   END_REGION

   REGION "CHANGE DETECTION"
       #old.btnParam := #btnParams;
       #old.kp8DI := #kp8DI;
       #old.logical := #retLogical.acutal;
       #old.physical := #btnPress;
   END_REGION

   REGION "OUTPUT"
       #kp8DQ := #colorMask;
       #physical := #retPhysical;
       #logical := #retLogical;
   END_REGION
END_FUNCTION_BLOCK

FUNCTION "KP8 Driver: HMI Emulator: Animation" : USInt   // FC26, SCL
{ S7_Optimized_Access := 'TRUE' }
VERSION : 0.1
   VAR_INPUT
      kp8Color : DWord;
      btnNumber : Int;
   END_VAR
   VAR_TEMP
      animate : USInt;
      blue : USInt;
      colorDWord : DWord;
      colorInt : DInt;
      green : USInt;
      off : USInt;
      red : USInt;
      white : USInt;
      yellow : USInt;
   END_VAR
   VAR CONSTANT
      blueMask : DInt := 16#0000_0100;
      btnMask : DInt := 16#0101_0100;
      greenMask : DInt := 16#0001_0000;
      offMask : DInt := 16#0000_0000;
      redMask : DInt := 16#0100_0000;
      whiteMask : DInt := 16#0101_0100;
      yellowMask : DInt := 16#0101_0000;
   END_VAR
BEGIN
   REGION "COPY TO LOCAL"
       #blue := "BLUE_LIGHT_BACKGROUND";
       #green := "GREEN_LIGHT_BACKGROUND";
       #off := "INVISIBLE";
       #red := "RED_LIGHT_BACKGROUND";
       #white := "WHITE_BACKGROUND";
       #yellow := "YELLOW_LIGHT_BACKGROUND";
   END_REGION

   REGION "ISOLATE BUTTON COLOR"
       #colorDWord := SHR_DWORD(IN := #kp8Color,N := INT_TO_ULINT(#btnNumber));
       #colorDWord := #colorDWord AND #btnMask;
       #colorInt := DWORD_TO_DINT(#colorDWord);
   END_REGION

   REGION "DETERMINE ANIMATION"
       CASE #colorInt OF
           #blueMask:
               #animate := #blue;
           #greenMask:
               #animate := #green;
           #redMask:
               #animate := #red;
           #whiteMask:
               #animate := #white;
           #yellowMask:
               #animate := #yellow;
           ELSE
               #animate := #off;
       END_CASE;
   END_REGION

   REGION "RETURN VALUE"
       #"KP8 Driver: HMI Emulator: Animation" := #animate;
   END_REGION
END_FUNCTION

FUNCTION "KP8 Driver: Group" : Void   // FC50, SCL
{ S7_Optimized_Access := 'TRUE' }
VERSION : 0.1
   VAR_INPUT
      btnNumber : Int;
      btnsParams : "KP8 Driver: Parameters: 8 Buttons";
   END_VAR
   VAR_IN_OUT
      logical : "KP8 Driver: Feedback Data";
   END_VAR
   VAR_TEMP
      pBtn : Int;
      retLogical : "KP8 Driver: Feedback Data";
      testGroup : Int;
      thisGroup : Int;
   END_VAR
BEGIN
   REGION "EXIT IF GROUP EQUALS 0"
       #thisGroup := #btnsParams.btn[#btnNumber].group;
       IF #thisGroup = 0 THEN
           RETURN;
       END_IF;
   END_REGION

   REGION "COPY TO LOCAL"
       #retLogical := #logical;
   END_REGION

   REGION "FOR EACH BUTTONS' PARAMETERS"
       FOR #pBtn := 0 TO 7 DO

           REGION "SKIP THE CURRENT BUTTON"
               IF #pBtn = #btnNumber THEN
                   GOTO NEXT;
               END_IF;
           END_REGION

           REGION "GROUP EXCLUSION"
               #testGroup := #btnsParams.btn[#pBtn].group;
               IF #testGroup = #thisGroup THEN
                   #retLogical.acutal.btn[#pBtn] := FALSE;
               END_IF;
           END_REGION

       NEXT:
           ;

       END_FOR;
   END_REGION

   REGION "OUTPUT"
       #logical := #retLogical;
   END_REGION
END_FUNCTION

FUNCTION "KP8 Driver: Toggle" : Void   // FC51, SCL
{ S7_Optimized_Access := 'TRUE' }
VERSION : 0.1
   VAR_INPUT
      signal : Bool;   // edge signal
   END_VAR
   VAR_IN_OUT
      state : Bool;   // logical button state
   END_VAR
BEGIN
   IF #signal THEN
       #state := NOT #state;
   END_IF;
END_FUNCTION

FUNCTION "KP8 Driver: Feedback" : Void   // FC52, SCL
{ S7_Optimized_Access := 'TRUE' }
VERSION : 0.1
   VAR_INPUT
      signal : Bool;
      oldSignal : Bool;
      btnNumber : Int;
   END_VAR
   VAR_IN_OUT
      feedback : "KP8 Driver: Feedback Data";
   END_VAR
   VAR_TEMP
      ret : "KP8 Driver: Feedback Data";
   END_VAR
BEGIN
   REGION "COPY TO LOCAL"
       #ret := #feedback;
       #ret.acutal.btn[#btnNumber] := #signal;
   END_REGION

   REGION "DEFAULT"
       #ret.rising.btn[#btnNumber] := FALSE;
       #ret.falling.btn[#btnNumber] := FALSE;
   END_REGION

   REGION "ON NEW INPUT"
       IF #signal <> #oldSignal THEN

           REGION "RISING EDGE"
               IF #signal AND NOT #oldSignal THEN
                   #ret.rising.btn[#btnNumber] := TRUE;
               END_IF;
           END_REGION

           REGION "FALLING EDGE"
               IF NOT #signal AND #oldSignal THEN
                   #ret.falling.btn[#btnNumber] := TRUE;
               END_IF;
           END_REGION

       END_IF;
   END_REGION


   REGION "OUTPUT"
       #feedback := #ret;
   END_REGION
END_FUNCTION

FUNCTION "KP8 Driver: State" : Void   // FC53, SCL
{ S7_Optimized_Access := 'TRUE' }
VERSION : 0.1
   VAR_INPUT
      press : "KP8 Driver: Feedback Data";
      btnNumber : Int;
      btnParams : "KP8 Driver: Parameters: 8 Buttons";
   END_VAR
   VAR_IN_OUT
      state : "KP8 Driver: Feedback Data";
   END_VAR
   VAR_TEMP
      pBtn : Int;
      retState : "KP8 Driver: Feedback Data";
   END_VAR
BEGIN
   REGION "RETURN ON INACTIVE BUTTON"
       IF NOT #btnParams.btn[#btnNumber].activate THEN
           RETURN;
       END_IF;
   END_REGION

   REGION "COPY TO LOCAL"
       #retState := #state;
   END_REGION

   REGION "MODE IS MOMENTARY"
       IF NOT #btnParams.btn[#btnNumber].mode THEN
           #retState.acutal.btn[#btnNumber] := #press.acutal.btn[#btnNumber];
       END_IF;
   END_REGION

   REGION "MAINTINED"
       IF #btnParams.btn[#btnNumber].mode THEN
           "KP8 Driver: Toggle"(signal := #press.rising.btn[#btnNumber],
                                state := #retState.acutal.btn[#btnNumber]);
       END_IF;
   END_REGION

   REGION "GROUP EXCLUSIVITY"
       IF #press.rising.btn[#btnNumber] THEN
           "KP8 Driver: Group"(btnNumber := #btnNumber,
                               btnsParams := #btnParams,
                               logical := #retState);
       END_IF;
   END_REGION

   REGION "OUTPUT"
       #state := #retState;
   END_REGION
END_FUNCTION

FUNCTION "KP8 Driver: Color" : Void   // FC54, SCL
{ S7_Optimized_Access := 'TRUE' }
VERSION : 0.1
   VAR_INPUT
      btnNum : Int;
      lblColor : String;   // 'red', 'green', 'blue', 'yellow', 'white', 'off'
   END_VAR
   VAR_IN_OUT
      btnColor : DWord;
   END_VAR
   VAR_TEMP
      btnMask : DWord;
      uColor : String;
      ret : DWord;
   END_VAR
   VAR CONSTANT
      btnMskRed : DWord := DWORD#16#0100_0000;
      btnMskGreen : DWord := DWORD#16#0001_0000;
      btnMskBlue : DWord := DWORD#16#0000_0100;
      btnMskYellow : DWord := DWORD#16#0101_0000;
      btnMskWhite : DWord := DWORD#16#0101_0100;
      btnMskOff : DWord := DWORD#16#FEFE_FEFF;
   END_VAR
BEGIN
   #ret := #btnColor;

   #ret := #ret AND ROL(IN := #btnMskOff,
                        N := INT_TO_UDINT(#btnNum));

   #uColor := #lblColor;
   "Upper"(#uColor);

   IF (#uColor = 'RED') THEN
       #btnMask := #btnMskRed;
   ELSIF (#uColor = 'GREEN') THEN
       #btnMask := #btnMskGreen;
   ELSIF (#uColor = 'BLUE') THEN
       #btnMask := #btnMskBlue;
   ELSIF (#uColor = 'YELLOW') THEN
       #btnMask := #btnMskYellow;
   ELSIF (#uColor = 'WHITE') THEN
       #btnMask := #btnMskWhite;
   ELSIF (#uColor = 'OFF') THEN
       ;
   END_IF;

   #ret := #ret OR SHL(IN := #btnMask,
                       N := INT_TO_UDINT(#btnNum));

   #btnColor := #ret;
END_FUNCTION

FUNCTION "KP8 Driver: HMI Emulator: Button Presses" : Word   // FC82, SCL
{ S7_Optimized_Access := 'TRUE' }
VERSION : 0.1
   VAR_INPUT
      pbs : DWord;
   END_VAR
   VAR_TEMP
      ret : Word;
   END_VAR
BEGIN
   #"KP8 Driver: HMI Emulator: Button Presses".%B1 := #pbs.%B0;
   #"KP8 Driver: HMI Emulator: Button Presses".%B0 := #pbs.%B1;
END_FUNCTION

// folder: Utilities

FUNCTION_BLOCK "Pulses: Button Collection"   // FB22, SCL
{ S7_Optimized_Access := 'TRUE' }
VERSION : 0.1
   VAR_INPUT
      btns : Variant;
   END_VAR
   VAR_IN_OUT
      pulses : Variant;
   END_VAR
   VAR
      old : Array[0..#u_bound] of Int;
   END_VAR
   VAR_TEMP
      eval : Array[0..#u_bound] of Int;
      i : Int;
      len_btns : UDInt;
      ret : Array[0..#u_bound] of Int;
      RET_VAL : Int;
   END_VAR
   VAR CONSTANT
      u_bound : Int := 999;
   END_VAR
BEGIN
   REGION "GET ARRAY LENGTH"
       #len_btns := CountOfElements(#btns);
   END_REGION


   REGION "COPY TO LOCAL"
       #RET_VAL := MOVE_BLK_VARIANT(SRC := #btns,
                                    COUNT := #len_btns,
                                    SRC_INDEX := 0,
                                    DEST_INDEX := 0,
                                    DEST => #eval);
   END_REGION


   REGION "CHECK FOR FALLING EDGE"
       FOR #i := 0 TO #u_bound DO
           IF #eval[#i] = 0 AND #old[#i] = 1 THEN
               #ret[#i] := 1;
           END_IF;
       END_FOR;
   END_REGION


   REGION "SAVE LAST SCAN"
       #old := #eval;
   END_REGION


   REGION "RETURN"
       #RET_VAL := MOVE_BLK_VARIANT(SRC := #ret,
                                    COUNT := #len_btns,
                                    SRC_INDEX := 0,
                                    DEST_INDEX := 0,
                                    DEST => #pulses);
   END_REGION
END_FUNCTION_BLOCK

FUNCTION_BLOCK "Push Button: State Changes"   // FB41, SCL
{ S7_Optimized_Access := 'TRUE' }
VERSION : 0.1
   VAR_IN_OUT
      interface : "Push Button Data";
      state_changes : "Push Button Data: State Change Data";
   END_VAR
   VAR
      old : "Push Button Data";
   END_VAR
   VAR_TEMP
      ret : Bool;
   END_VAR
BEGIN
   REGION "ACTUATE"
       #state_changes.actuate.actual := #interface.actuate;
       #state_changes.actuate.rising := "Bool.Rising_Edge"(signal := #interface.actuate,
                                                            old_signal := #old.actuate);
       #state_changes.actuate.falling := "Bool.Falling_Edge"(signal := #interface.actuate,
                                                              old_signal := #old.actuate);
   END_REGION

   REGION "ANIMATE"
       #state_changes.animate.rising := "USInt.Value_Change"(value := #interface.animate,
                                                         old_value := #old.animate);
       #state_changes.animate.actual := #interface.animate;
       #state_changes.animate.falling := FALSE;     // animate never set to null token
   END_REGION

   REGION "ENABLE"
       #state_changes.enable.rising := "Bool.Rising_Edge"(signal := #interface.enable,
                                                           old_signal := #old.enable);
       #state_changes.enable.actual := #interface.enable;
       #state_changes.enable.falling := "Bool.Falling_Edge"(signal := #interface.enable,
                                                             old_signal := #old.enable);
   END_REGION

   REGION "LABEL"
       #state_changes.label.rising := "WString: Rising Edge"(value := #interface.label,
                                                        old_value := #old.label);
       #state_changes.label.actual := #interface.label;
       #state_changes.label.falling := "WString: Falling Edge"(value := #interface.label,
                                                          old_value := #old.label);
   END_REGION

   REGION "LIST SELECT"
       #state_changes.listSelect.rising := "UInt.Value_Change"(value := #interface.listSelect,
                                                           old_value := #old.listSelect);
       #state_changes.listSelect.actual := #interface.listSelect;
       #state_changes.listSelect.falling := FALSE;      // list select never set to null token
   END_REGION

   REGION "VISIBLE"
       #state_changes.visible.rising := "Bool.Rising_Edge"(signal := #interface.visible,
                                                       old_signal := #old.visible);
       #state_changes.visible.actual := #interface.visible;
       #state_changes.visible.falling := "Bool.Falling_Edge"(signal := #interface.visible,
                                                         old_signal := #old.visible);
   END_REGION

   REGION "SAVE OLD VALUES"
       #old := #interface;
   END_REGION
END_FUNCTION_BLOCK

FUNCTION_BLOCK "IO Field: State Changes"   // FB48, SCL
{ S7_Optimized_Access := 'TRUE' }
VERSION : 0.1
   VAR_IN_OUT
      interface : "IO Field Data: Label with Data";
      feedback : "IO Field: State Change Data";
   END_VAR
   VAR
      old : "IO Field Data: Label with Data";
   END_VAR
BEGIN
   REGION "ANIMATE"
       #feedback.animate.rising := "USInt.Value_Change"(value := #interface.animate,
                                                         old_value := #old.animate);
       #feedback.animate.actual := #interface.animate;
       #feedback.animate.falling := FALSE;     // animate never set to null token 
   END_REGION

   REGION "ENABLE"
       #feedback.enable.rising := "Bool.Rising_Edge"(signal := #interface.enable,
                                                      old_signal := #old.enable);
       #feedback.enable.actual := #interface.enable;
       #feedback.enable.falling := "Bool.Falling_Edge"(signal := #interface.enable,
                                                        old_signal := #old.enable);
   END_REGION

   REGION "INPUT FINISHED"
       #feedback.input_finished.rising := "Bool.Rising_Edge"(signal := #interface.input_finished,
                                                              old_signal := #old.input_finished);
       #feedback.input_finished.actual := #interface.input_finished;
       #feedback.input_finished.falling := "Bool.Falling_Edge"(signal := #interface.input_finished,
                                                                old_signal := #old.input_finished);
   END_REGION

   REGION "VALUE CHANGED"
       #feedback.value.rising := "WString: Rising Edge"(value := #interface.value,
                                                        old_value := #old.value);
       #feedback.value.actual := #interface.value;
       #feedback.value.falling := "WString: Falling Edge"(value := #interface.value,
                                                          old_value := #old.value);
   END_REGION

   REGION "VISIBLE"
       #feedback.visible.rising := "Bool.Rising_Edge"(signal := #interface.visible,
                                                       old_signal := #old.visible);
       #feedback.visible.actual := #interface.visible;
       #feedback.visible.falling := "Bool.Falling_Edge"(signal := #interface.visible,
                                                         old_signal := #old.visible);
   END_REGION

   REGION "SAVE OLD VALUES"
       #old := #interface;
   END_REGION
END_FUNCTION_BLOCK

FUNCTION_BLOCK "Get Data: WString"   // FB51, SCL
{ S7_Optimized_Access := 'TRUE' }
VERSION : 0.1
   VAR_INPUT
      value : WString;
   END_VAR
   VAR_IN_OUT
      get_wstring : "State Changes: WString";
   END_VAR
   VAR
      old_value : WString;
   END_VAR
   VAR_TEMP
      ret : "State Changes: WString";
   END_VAR
   VAR CONSTANT
      blank : WString;
   END_VAR
BEGIN
   REGION "BUFFER IN"
       #ret := #get_wstring;
   END_REGION

   REGION "MAP"
       IF #value <> #old_value THEN
           #get_wstring.actual := #value;
       END_IF;
       #ret.rising := "WString: Rising Edge"(value := #value, old_value := #old_value);
       #ret.falling := "WString: Falling Edge"(value := #value, old_value := #old_value);
   END_REGION

   REGION "SAVE OLD VALUE"
       #old_value := #value;
   END_REGION


   REGION "RETURN" 
       #get_wstring := #ret;
   END_REGION
END_FUNCTION_BLOCK

FUNCTION_BLOCK "Get Data: Real"   // FB52, SCL
{ S7_Optimized_Access := 'TRUE' }
VERSION : 0.1
   VAR_INPUT
      value : WString;
   END_VAR
   VAR_IN_OUT
      get_real : "State Changes: Real";
   END_VAR
   VAR
      old_value : WString;
   END_VAR
   VAR_TEMP
      ret : "State Changes: Real";
   END_VAR
   VAR CONSTANT
      blank : WString;
   END_VAR
BEGIN
   REGION "BUFFER IN"
       #ret := #get_real;
   END_REGION

   REGION "MAP"
       IF #value <> #old_value THEN
           #get_real.actual := "Timer.WString_to_Real"(#value);
       END_IF;
       #ret.rising := "WString: Rising Edge"(value := #value, old_value := #old_value);
       #ret.falling := "WString: Falling Edge"(value := #value, old_value := #old_value);
   END_REGION

   REGION "SAVE OLD VALUE"
       #old_value := #value;
   END_REGION


   REGION "RETURN" 
       #get_real := #ret;
   END_REGION
END_FUNCTION_BLOCK

FUNCTION "Pointer Calc: KP8 Labels" : Int   // FC25, SCL
{ S7_Optimized_Access := 'TRUE' }
VERSION : 0.1
   VAR_INPUT
      index : Int;
   END_VAR
   VAR_TEMP
      val : Int;
   END_VAR
BEGIN
   IF #index >= 4 THEN
       #val := 7 - (#index - 4) * 2;
   END_IF;

   IF #index <= 3 THEN
       #val := 8 - #index * 2;
   END_IF;

   #"Pointer Calc: KP8 Labels" := #val;
END_FUNCTION

FUNCTION "Row Pointer: Roll Over" : Void   // FC33, SCL
{ S7_Optimized_Access := 'TRUE' }
VERSION : 0.1
   VAR_INPUT
      limit : Int;
   END_VAR
   VAR_IN_OUT
      pointer : Int;
   END_VAR
BEGIN
   REGION "INCREMENT"
       #pointer += 1;
   END_REGION

   REGION "HIGH LIMIT ROLLOVER"
       IF #pointer > "partReqDataRowCount" THEN
           #pointer := 0;
       END_IF;
   END_REGION
END_FUNCTION

FUNCTION "KP8.DURL_to_LRUD" : Int   // FC35, SCL
{ S7_Optimized_Access := 'TRUE' }
VERSION : 0.1
   VAR_INPUT
      btnNum : Int;
   END_VAR
   VAR_TEMP
      output : Int;
   END_VAR
BEGIN
   IF #btnNum MOD 2 = 0 THEN
       #output := 7 - #btnNum / 2;
   END_IF;
   IF #btnNum MOD 2 <> 0 THEN
       #output := 3 - #btnNum / 2;
   END_IF;
   #"KP8.DURL_to_LRUD" := #output;
END_FUNCTION

FUNCTION "Validate PN" : Bool   // FC42, SCL
{ S7_Optimized_Access := 'TRUE' }
VERSION : 0.1
   VAR_INPUT
      pnCode : DInt;
      pnLib : "Recipe: PN Text Library";
   END_VAR
   VAR_TEMP
      pn : WString;
      ret : Bool;
   END_VAR
BEGIN
   REGION "GET PN FROM LIBRARY"
       #pn := "Part_Number.Code_to_WString"(pnLib := #pnLib,
                                pnCode := #pnCode);
   END_REGION

   REGION "BUTTON HAS NO PN"
       IF LEN(#pn) = 0 THEN
           #ret := FALSE;
       END_IF;
   END_REGION

   REGION "BUTTON HAS PN"
       IF LEN(#pn) <> 0 THEN
           #ret := TRUE;
       END_IF;
   END_REGION

   REGION "RETURN"
       #"Validate PN" := #ret;
   END_REGION
END_FUNCTION

FUNCTION "Row Pointer: Post Collapse" : Void   // FC56, SCL
{ S7_Optimized_Access := 'TRUE' }
VERSION : 0.1
   VAR_INPUT
      dataTable : "Part Request Data";
   END_VAR
   VAR_IN_OUT
      pDataRow : Int;
   END_VAR
   VAR_TEMP
      pRow : Int;
   END_VAR
BEGIN
   REGION "SCAN TABLE"
       WHILE #dataTable.row[#pRow] <> -1 AND #pRow <= "partReqDataRowCount" DO
           #pRow += 1;
       END_WHILE;
   END_REGION

   REGION "TABLE NOT FULL"
       IF #pRow <="partReqDataRowCount" THEN
           #pDataRow := #pRow;
           RETURN;
       END_IF;
   END_REGION

   REGION "TABLE FULL"
       IF #pRow > "partReqDataRowCount" THEN
           #pDataRow := 0;
           RETURN;
       END_IF;
   END_REGION
END_FUNCTION

FUNCTION "Part Ordered" : Bool   // FC90, SCL
{ S7_Optimized_Access := 'TRUE' }
VERSION : 0.1
// checks state to see if the part has been ordered by the warehouse; returns a bool
   VAR_INPUT
      state : Int;
   END_VAR
   VAR_TEMP
      ret : Bool;
   END_VAR
BEGIN
   IF #state / 10 = 2 THEN
       #ret := TRUE;
   END_IF;
   #"Part Ordered" := #ret;
END_FUNCTION

FUNCTION "Is_HMI_Station" : Bool   // FC96, SCL
{ S7_Optimized_Access := 'TRUE' }
VERSION : 0.1
   VAR_INPUT
      stn : "Station: Single Station";
   END_VAR
   VAR_TEMP
      ret : Bool;
   END_VAR
BEGIN
   REGION "CHECK WIP COUNT"
       IF #stn.wipData.count > 0 THEN
           #ret := TRUE;
       END_IF;
   END_REGION


   REGION "RETURN"
       #Is_HMI_Station := #ret;
   END_REGION
END_FUNCTION

FUNCTION "Toggle" : Void   // FC103, SCL
{ S7_Optimized_Access := 'TRUE' }
VERSION : 0.1
   VAR_INPUT
      pulse : Bool;
   END_VAR
   VAR_IN_OUT
      state : Bool;
   END_VAR
   VAR_TEMP
      ret : Bool;
   END_VAR
BEGIN
   REGION "COPY TO LOCAL"
       #ret := #state;
   END_REGION


   REGION "TOGGLE ON PULSE"
       IF #pulse THEN
           #ret := NOT #ret;
       END_IF;
   END_REGION


   REGION "RETURN"
       #state := #ret;
   END_REGION
END_FUNCTION

FUNCTION "Count Selected Stations" : Int   // FC105, SCL
{ S7_Optimized_Access := 'TRUE' }
VERSION : 0.1
   VAR_INPUT
      selected_stns : Array[0.."STATION_COUNT"] of Bool;
   END_VAR
   VAR_TEMP
      count : Int;
      i : Int;
   END_VAR
BEGIN
   REGION "CHECK EACH STATION"
       FOR #i := 0 TO "STATION_COUNT" DO
           IF #selected_stns[#i] THEN
               #count += 1;
           END_IF;
       END_FOR;
   END_REGION


   REGION "RETURN COUNT"
       #"Count Selected Stations" := #count;
   END_REGION
END_FUNCTION

FUNCTION "Get Station Index From Id" : Int   // FC106, SCL
{ S7_Optimized_Access := 'TRUE' }
VERSION : 0.1
   VAR_INPUT
      line_name : WString;
      drop_zone : USInt;
      stns : "Station: All Stations";
   END_VAR
   VAR_TEMP
      i : Int;
      ret : Int;
   END_VAR
BEGIN
   REGION "MATCH LINE NAME AND DROP ZONE"
       FOR #i := 0 TO "STATION_COUNT" DO
           IF #line_name = #stns.stn[#i].id.lineName THEN
               IF #drop_zone = #stns.stn[#i].id.dropZone THEN
                   #ret := #i;
                   EXIT;
               END_IF;
           END_IF;
       END_FOR;
   END_REGION


   REGION "RETURN"
       #"Get Station Index From Id" := #ret;
   END_REGION
END_FUNCTION

FUNCTION "Get First Selected Station" : Int   // FC108, SCL
{ S7_Optimized_Access := 'TRUE' }
VERSION : 0.1
   VAR_INPUT
      selected_stns : Array[0.."STATION_COUNT"] of Bool;
   END_VAR
   VAR_TEMP
      eval_station_index : Int;
      i : Int;
   END_VAR
BEGIN
   REGION "FIND FIRST SELECTED STATION"
       FOR #i := 0 TO "STATION_COUNT" DO
           IF #selected_stns[#i] THEN
               #eval_station_index := #i;
               EXIT;
           END_IF;
       END_FOR;
   END_REGION


   REGION "RETURN"
       #"Get First Selected Station" := #eval_station_index;
   END_REGION
END_FUNCTION

FUNCTION "Remap Int Array" : Void   // FC122, SCL
{ S7_Optimized_Access := 'TRUE' }
VERSION : 0.1
   VAR_INPUT
      source_int_array : Variant;
   END_VAR
   VAR_IN_OUT
      destination_int_array : Variant;
   END_VAR
   VAR_TEMP
      len_destination : UDInt;
      status : Int;
   END_VAR
BEGIN
   #len_destination := CountOfElements(#destination_int_array);
   #status := MOVE_BLK_VARIANT(SRC := #source_int_array,
                               COUNT := #len_destination,
                               SRC_INDEX := 0,
                               DEST_INDEX := 0,
                               DEST => #destination_int_array);
END_FUNCTION

FUNCTION "Count Selected WIPs" : Int   // FC126, SCL
{ S7_Optimized_Access := 'TRUE' }
VERSION : 0.1
   VAR_INPUT
      selected_WIPs : Array[0.."WIP_COUNT"] of DInt;
   END_VAR
   VAR_TEMP
      count : Int;
      i : Int;
   END_VAR
BEGIN
   REGION "CHECK EACH STATION"
       FOR #i := 0 TO "WIP_COUNT" DO
           IF #selected_WIPs[#i] = INT_TO_DINT("NULL_TOKEN") THEN
               EXIT;
           END_IF;
           IF #selected_WIPs[#i] <> INT_TO_DINT("NULL_TOKEN") THEN
               #count += 1;
           END_IF;
       END_FOR;
   END_REGION


   REGION "RETURN COUNT"
       #"Count Selected WIPs" := #count;
   END_REGION
END_FUNCTION

FUNCTION "Count Selected Buttons" : Int   // FC127, SCL
{ S7_Optimized_Access := 'TRUE' }
VERSION : 0.1
   VAR_INPUT
      selected_buttons : Array[0.."STATION_BUTTON_COUNT"] of Bool;
   END_VAR
   VAR_TEMP
      count : Int;
      i : Int;
   END_VAR
BEGIN
   REGION "CHECK EACH STATION"
       FOR #i := 0 TO "STATION_BUTTON_COUNT" DO
           IF #selected_buttons[#i] THEN
               #count += 1;
           END_IF;
       END_FOR;
   END_REGION


   REGION "RETURN COUNT"
       #"Count Selected Buttons" := #count;
   END_REGION
END_FUNCTION

FUNCTION "Collapse DInt Array" : Void   // FC132, SCL
{ S7_Optimized_Access := 'TRUE' }
VERSION : 0.1
   VAR_INPUT
      null_value : DInt;   // value that indicates null data
   END_VAR
   VAR_IN_OUT
      int_array : Variant;
   END_VAR
   VAR_TEMP
      i : Int;
      j : Int;
      len_int : Int;
      len_udint : UDInt;
      status : Int;
      t_int_array : Array[0..999] of DInt;
   END_VAR
BEGIN
   REGION "COPY TO LOCAL MEMORY"
       #len_udint := CountOfElements(#int_array);
       #len_int := UDINT_TO_INT(#len_udint) - 1;
       #status := MOVE_BLK_VARIANT(SRC := #int_array,
                                   COUNT := #len_udint,
                                   SRC_INDEX := 0,
                                   DEST_INDEX := 0,
                                   DEST => #t_int_array);
   END_REGION

   REGION "COLLAPSE IN PLACE"
       FOR #i := 0 TO #len_int - 1 DO
           IF #t_int_array[#i] = #null_value THEN
               FOR #j := #i + 1 TO #len_int DO
                   IF #t_int_array[#j] <> #null_value THEN
                       #t_int_array[#i] := #t_int_array[#j];
                       #t_int_array[#j] := #null_value;
                       EXIT;
                   END_IF;
               END_FOR;
           END_IF;
       END_FOR;
   END_REGION

   REGION "RETURN"
       #status := MOVE_BLK_VARIANT(SRC := #t_int_array,
                                   COUNT := #len_udint,
                                   SRC_INDEX := 0,
                                   DEST_INDEX := 0,
                                   DEST => #int_array);
   END_REGION
END_FUNCTION

FUNCTION "Count Collapsed DInt Array" : Int   // FC133, SCL
{ S7_Optimized_Access := 'TRUE' }
VERSION : 0.1
   VAR_INPUT
      null_value : DInt;
      "array" : Variant;
   END_VAR
   VAR_TEMP
      count : Int;
      i : Int;
      len_int : Int;
      len_udint : UDInt;
      status : Int;
      t_array : Array[0..999] of DInt;
   END_VAR
BEGIN
   REGION "NOTES"
       (*
       returns the number of valid elements in a collapsed int array
       *)
   END_REGION


   REGION "COPY TO LOCAL"
       #len_udint := CountOfElements(#array);
       #len_int := UDINT_TO_INT(#len_udint) - 1;
       #status := MOVE_BLK_VARIANT(SRC := #array,
                                   COUNT := #len_udint,
                                   SRC_INDEX := 0,
                                   DEST_INDEX := 0,
                                   DEST => #t_array);
   END_REGION


   REGION "SCAN FOR FIRST NULL"
       FOR #i := 0 TO #len_int DO
           IF #t_array[#i] = INT_TO_DINT("NULL_TOKEN") THEN
               EXIT;
           END_IF;
           IF #t_array[#i] <> #null_value THEN
               #count += 1;
           END_IF;
       END_FOR;
   END_REGION


   REGION "RETURN"
       #"Count Collapsed DInt Array" := #count;
   END_REGION
END_FUNCTION

FUNCTION "Map WIP Codes to DInt Array" : Void   // FC139, SCL
{ S7_Optimized_Access := 'TRUE' }
VERSION : 0.1
   VAR_INPUT
      station : "WIP: Station";
   END_VAR
   VAR_IN_OUT
      WIP_array : Array[0.."WIP_COUNT"] of DInt;
   END_VAR
   VAR_TEMP
      i : Int;
   END_VAR
BEGIN
   FOR #i := 0 TO "WIP_COUNT" DO
       IF #station.wip[#i].wip.code = "NULL_TOKEN" THEN
           EXIT;
       END_IF;
       #WIP_array[#i] := #station.wip[#i].wip.code;
   END_FOR;
END_FUNCTION

FUNCTION "Map Selected Stations to Int Array" : Void   // FC142, SCL
{ S7_Optimized_Access := 'TRUE' }
VERSION : 0.1
   VAR_INPUT
      selected_stations : "Selected Stations";
   END_VAR
   VAR_OUTPUT
      selected_stations_indicies : Array[0.."STATION_COUNT"] of Int;
   END_VAR
   VAR_TEMP
      i : Int;
      p_ret : Int;
      _return : Array[0.."STATION_COUNT"] of Int;
   END_VAR
BEGIN
   "Array.Int.Fill"(value := "NULL_TOKEN",
                    int_array := #_return);
   FOR #i := 0 TO "STATION_COUNT" DO
       IF #selected_stations.stns[#i] THEN
           #_return[#p_ret] := #i;
           #p_ret += 1;
       END_IF;
   END_FOR;
   #selected_stations_indicies := #_return;
END_FUNCTION

FUNCTION "USInt.Value_Change" : Bool   // FC181, SCL
{ S7_Optimized_Access := 'TRUE' }
VERSION : 0.1
   VAR_INPUT
      value : USInt;
      old_value : USInt;
   END_VAR
BEGIN
   #"USInt.Value_Change" := #value <> #old_value;
END_FUNCTION

// folder: Utilities/Address

FUNCTION "Address.Get_Button" : DInt   // FC21, SCL
{ S7_Optimized_Access := 'TRUE' }
VERSION : 0.1
   VAR_INPUT
      address : DInt;
   END_VAR
BEGIN
   #"Address.Get_Button" := #address MOD 10;
END_FUNCTION

FUNCTION "Address.Get_Station" : DInt   // FC24, SCL
{ S7_Optimized_Access := 'TRUE' }
VERSION : 0.1
   VAR_INPUT
      address : DInt;
   END_VAR
BEGIN
   #"Address.Get_Station" := #address / 10_000;
END_FUNCTION

FUNCTION "Address.Set_Address" : DInt   // FC32, SCL
{ S7_Optimized_Access := 'TRUE' }
VERSION : 0.1
   VAR_INPUT
      pBtn : Int;
      pStn : Int;
      pWip : Int;
   END_VAR
BEGIN
   #"Address.Set_Address" := INT_TO_DINT(#pStn) * 10_000 + INT_TO_DINT(#pWip) * 10 + INT_TO_DINT(#pBtn);
END_FUNCTION

FUNCTION "Address.Get_Wip" : DInt   // FC88, SCL
{ S7_Optimized_Access := 'TRUE' }
VERSION : 0.1
   VAR_INPUT
      address : DInt;
   END_VAR
BEGIN
   #"Address.Get_Wip" := #address - "Address.Get_Station"(#address) * 10_000 - "Address.Get_Button"(#address);
END_FUNCTION

// folder: Utilities/Array

FUNCTION "Array.Any.Length" : UDInt   // FC60, SCL
{ S7_Optimized_Access := 'TRUE' }
VERSION : 0.1
   VAR_INPUT
      "array" : Variant;
   END_VAR
   VAR_TEMP
      status : DInt;
      ret : UDInt;
   END_VAR
BEGIN
   #ret := CountOfElements(#array);
   #"Array.Any.Length" := #ret;
END_FUNCTION

FUNCTION "Array.Int.Fill" : Void   // FC109, SCL
{ S7_Optimized_Access := 'TRUE' }
VERSION : 0.1
   VAR_INPUT
      value : Int;
   END_VAR
   VAR_IN_OUT
      int_array : Array[*] of Int;
   END_VAR
   VAR_TEMP
      _i : DInt;
      _length : DInt;
   END_VAR
BEGIN
   REGION "GET LENGHT"
       #_length := UDINT_TO_DINT("Array.Any.Length"(#int_array));
       #_length -= 1;
   END_REGION


   REGION "FILL LENGTH WITH BYTE IN"
       FOR #_i := 0 TO #_length DO
           #int_array[#_i] := #value;
       END_FOR;
   END_REGION
END_FUNCTION

FUNCTION "Array.DInt.Is_Element" : Bool   // FC111, SCL
{ S7_Optimized_Access := 'TRUE' }
VERSION : 0.1
   VAR_INPUT
      dint_array : Array[*] of DInt;
      search_term : DInt;
   END_VAR
   VAR_TEMP
      _i : DInt;
      _length : DInt;
   END_VAR
BEGIN
   REGION "LOCAL VARIABLES"
       #_length := UDINT_TO_DINT("Array.Any.Length"(#dint_array)) - 1;
   END_REGION


   REGION "SEARCH ARRAY"
       FOR #_i := 0 TO #_length DO
           IF #dint_array[#_i] <> #search_term THEN
               CONTINUE;
           END_IF;
           #"Array.DInt.Is_Element" := TRUE;
           RETURN;
       END_FOR;
   END_REGION


   REGION "NOT FOUND"
       #"Array.DInt.Is_Element" := FALSE;
       RETURN;
   END_REGION
END_FUNCTION

FUNCTION "Array.Int.Collapse" : Void   // FC114, SCL
{ S7_Optimized_Access := 'TRUE' }
VERSION : 0.1
   VAR_INPUT
      null_value : Int;   // value that indicates null data
   END_VAR
   VAR_IN_OUT
      int_array : Variant;
   END_VAR
   VAR_TEMP
      i : Int;
      j : Int;
      len_int : Int;
      len_udint : UDInt;
      status : Int;
      t_int_array : Array[0..999] of Int;
   END_VAR
BEGIN
   REGION "COPY TO LOCAL MEMORY"
       #len_udint := CountOfElements(#int_array);
       #len_int := UDINT_TO_INT(#len_udint) - 1;
       #status := MOVE_BLK_VARIANT(SRC := #int_array,
                                   COUNT := #len_udint,
                                   SRC_INDEX := 0,
                                   DEST_INDEX := 0,
                                   DEST => #t_int_array);
   END_REGION

   REGION "COLLAPSE IN PLACE"
       FOR #i := 0 TO #len_int - 1 DO
           IF #t_int_array[#i] = #null_value THEN
               FOR #j := #i + 1 TO #len_int DO
                   IF #t_int_array[#j] <> #null_value THEN
                       #t_int_array[#i] := #t_int_array[#j];
                       #t_int_array[#j] := #null_value;
                       EXIT;
                   END_IF;
               END_FOR;
           END_IF;
       END_FOR;
   END_REGION

   REGION "RETURN"
       #status := MOVE_BLK_VARIANT(SRC := #t_int_array,
                                   COUNT := #len_udint,
                                   SRC_INDEX := 0,
                                   DEST_INDEX := 0,
                                   DEST => #int_array);
   END_REGION
END_FUNCTION

FUNCTION "Array.Int.Count" : Int   // FC115, SCL
{ S7_Optimized_Access := 'TRUE' }
VERSION : 0.1
   VAR_INPUT
      null_value : Int;
      "array" : Variant;
   END_VAR
   VAR_TEMP
      count : Int;
      i : Int;
      len_int : Int;
      len_udint : UDInt;
      status : Int;
      t_array : Array[0..999] of Int;
   END_VAR
BEGIN
   REGION "NOTES"
       (*
       returns the number of valid elements in a collapsed int array
       *)
   END_REGION


   REGION "COPY TO LOCAL"
       #len_udint := CountOfElements(#array);
       #len_int := UDINT_TO_INT(#len_udint) - 1;
       #status := MOVE_BLK_VARIANT(SRC := #array,
                                   COUNT := #len_udint,
                                   SRC_INDEX := 0,
                                   DEST_INDEX := 0,
                                   DEST => #t_array);
   END_REGION


   REGION "SCAN FOR FIRST NULL"
       FOR #i := 0 TO #len_int DO
           IF #t_array[#i] = #null_value THEN
               EXIT;
           END_IF;
           IF #t_array[#i] <> #null_value THEN
               #count += 1;
           END_IF;
       END_FOR;
   END_REGION


   REGION "RETURN"
       #"Array.Int.Count" := #count;
   END_REGION
END_FUNCTION

FUNCTION "Array.Bool.True_Indices" : Void   // FC120, SCL
{ S7_Optimized_Access := 'TRUE' }
VERSION : 0.1
   VAR_INPUT
      array_of_bool : Array[*] of Bool;   // max 1000 elements
   END_VAR
   VAR_IN_OUT
      list_of_indices : Array[*] of Int;   // max 1000 elements
   END_VAR
   VAR_TEMP
      _i : Int;
      _length : Int;
      _p_return : Int;
      _resized_bool_array : Array[0..#UBOUND] of Bool;
   END_VAR
   VAR CONSTANT
      UBOUND : Int := 999;
   END_VAR
BEGIN
   REGION "FILL RETURN ARRAY"
       "Array.Int.Fill"(value := "NULL_TOKEN",
                        int_array := #list_of_indices);
   END_REGION


   REGION "COPY TO ARRAY OF STATIC SIZE"
       #_length := UDINT_TO_INT("Array.Any.Length"(#array_of_bool)) - 1;
       FOR #_i := 0 TO #_length DO
           #_resized_bool_array[#_i] := #array_of_bool[#_i];
       END_FOR;
   END_REGION


   REGION "INSERT INDICES INTO RETURN ARRAY"
       FOR #_i := 0 TO #UBOUND DO
           IF #_resized_bool_array[#_i] THEN
               #list_of_indices[#_p_return] := #_i;
               #_p_return += 1;
           END_IF;
       END_FOR;
   END_REGION
END_FUNCTION

FUNCTION "Array.Int.Is_Element" : Bool   // FC121, SCL
{ S7_Optimized_Access := 'TRUE' }
VERSION : 0.1
   VAR_INPUT
      int_array : Array[*] of Int;
      search_term : Int;
   END_VAR
   VAR_TEMP
      _i : Int;
      _length : DInt;
   END_VAR
BEGIN
   REGION "LOCAL VARIABLES"
       #_length := UDINT_TO_DINT("Array.Any.Length"(#int_array)) - 1;
   END_REGION


   REGION "SEARCH ARRAY"
       FOR #_i := 0 TO #_length DO
           IF #int_array[#_i] <> #search_term THEN
               CONTINUE;
           END_IF;
           #"Array.Int.Is_Element" := TRUE;
           RETURN;
       END_FOR;
   END_REGION


   REGION "NOT FOUND"
       #"Array.Int.Is_Element" := FALSE;
       RETURN;
   END_REGION
END_FUNCTION

FUNCTION "Array.DInt.Fill" : Void   // FC131, SCL
{ S7_Optimized_Access := 'TRUE' }
VERSION : 0.1
   VAR_INPUT
      int_in : DInt;
   END_VAR
   VAR_OUTPUT
      array_out : Variant;
   END_VAR
   VAR_TEMP
      i : Int;
      internal_array : Array[0..999] of DInt;
      len_array_out : UDInt;
      status : Int;
   END_VAR
BEGIN
   REGION "GET LENGHT"
       #len_array_out := CountOfElements(#array_out);
   END_REGION


   REGION "FILL LENGTH WITH BYTE IN"
       FOR #i := 0 TO UDINT_TO_INT(#len_array_out) - 1 DO
           #internal_array[#i] := #int_in;
       END_FOR;
   END_REGION


   REGION "RETURN"
       #status := MOVE_BLK_VARIANT(SRC := #internal_array,
                                   COUNT := #len_array_out,
                                   SRC_INDEX := 0,
                                   DEST_INDEX := 0,
                                   DEST => #array_out);
   END_REGION
END_FUNCTION

FUNCTION "Array.Int.Search" : Int   // FC140, SCL
{ S7_Optimized_Access := 'TRUE' }
VERSION : 0.1
   VAR_INPUT
      array_of_int : Variant;   // max upper bound 999
      search_term : Int;
   END_VAR
   VAR_TEMP
      i : Int;
      len_as_udint : UDInt;
      len_as_int : Int;
      ret : Int;
      status : Int;
      t_array : Array[0..999] of Int;
   END_VAR
   // Ret_Val : index of search term. returns -1 if not found.
BEGIN
   REGION "LOCAL VARIABLES"
       #len_as_udint := CountOfElements(#array_of_int);
       #len_as_int := UDINT_TO_INT(#len_as_udint) - 1;
       #status := MOVE_BLK_VARIANT(SRC := #array_of_int,
                                   COUNT := #len_as_udint,
                                   SRC_INDEX := 0,
                                   DEST_INDEX := 0,
                                   DEST => #t_array);
       #ret := -1;
   END_REGION


   REGION "SEARCH ARRAY"
       FOR #i := 0 TO #len_as_int DO
           IF #t_array[#i] = #search_term THEN
               #ret := #i;
               EXIT;
           END_IF;
       END_FOR;
   END_REGION


   REGION "RETURN"
       #"Array.Int.Search" := #ret;
   END_REGION
END_FUNCTION

FUNCTION "Array.Int.Intersect" : Void   // FC141, SCL
{ S7_Optimized_Access := 'TRUE' }
VERSION : 0.1
   VAR_INPUT
      "a" : Variant;   // should be array of int, max 999
      "b" : Variant;   // should be array of int, max 999
      null_value : Int;
   END_VAR
   VAR_OUTPUT
      intersect_array : Variant;   // should be array of int, max 999
   END_VAR
   VAR_TEMP
      i : Int;
      j : Int;
      len_a : Struct
         as_udint : UDInt;
         as_int : Int;
      END_STRUCT;
      len_b : Struct
         as_udint : UDInt;
         as_int : Int;
      END_STRUCT;
      len_longer : Struct
         as_udint : UDInt;
         as_int : Int;
      END_STRUCT;
      len_shorter : Struct
         as_udint : UDInt;
         as_int : Int;
      END_STRUCT;
      t_a : Array[0..#u_bound] of Int;
      p_ret : Int;
      ret : Array[0..#u_bound_double] of Int;
      t_b : Array[0..#u_bound] of Int;
      status : Int;
   END_VAR
   VAR CONSTANT
      u_bound : Int := 999;
      u_bound_double : Int := 1999;
   END_VAR
BEGIN
   REGION "GET LENGTHS"
       #len_a.as_udint := CountOfElements(#a);
       #len_a.as_int := UDINT_TO_INT(#len_a.as_udint) - 1;
       #len_b.as_udint := CountOfElements(#b);
       #len_b.as_int := UDINT_TO_INT(#len_b.as_udint) - 1;
   END_REGION

   REGION "MOVE"
       #status := MOVE_BLK_VARIANT(SRC := #a, COUNT := #len_a.as_udint, SRC_INDEX := 0, DEST_INDEX := 0, DEST => #t_a);
       #status := MOVE_BLK_VARIANT(SRC := #b, COUNT := #len_b.as_udint, SRC_INDEX := 0, DEST_INDEX := 0, DEST => #t_b);
   END_REGION

   REGION "FIND INTERSECT"
       FOR #i := 0 TO #len_a.as_int DO
           IF #t_a[#i] = #null_value THEN
               EXIT;
           END_IF;
           FOR #j := 0 TO #len_b.as_int DO
               IF #t_b[#j] = #null_value THEN
                   EXIT;
               END_IF;
               IF #t_a[#i] = #t_b[#j] THEN
                   #ret[#p_ret] := #t_a[#i];
                   #p_ret += 1;
                   EXIT;
               END_IF;
           END_FOR;
       END_FOR;
   END_REGION

   REGION "RETURN"
       #status := MOVE_BLK_VARIANT(SRC := #ret, COUNT := INT_TO_UDINT(#p_ret - 1), SRC_INDEX := 0, DEST_INDEX := 0, DEST => #intersect_array);
   END_REGION
END_FUNCTION

FUNCTION "Array.DInt.First_Occurance" : DInt   // FC143, SCL
{ S7_Optimized_Access := 'TRUE' }
VERSION : 0.1
   VAR_INPUT
      dint_array : Array[*] of DInt;
      search_term : Int;
   END_VAR
   VAR_TEMP
      _i : DInt;
      _length : UDInt;
   END_VAR
BEGIN
   REGION "NOTES"
       (* 
       This function returns the first occurance of the search term.
       This function meant for use with collapsed arrays.
       See "Array.DInt.Collapse" for collapse functionality.
       *)
   END_REGION


   REGION "GET LENGTH OF INPUT ARRAY"
       #_length := "Array.Any.Length"(#dint_array);
   END_REGION


   REGION "FIND FIRST SEARCH TERM, -1 IF NONE"
       (*
       Its worth noting that "Array.DInt.Is_Element" could return the index of the search term
       as an output, saving the processor some work. 
       The rework is justified by increased encapsulation.
       The time complexity for "Array.DInt.First_Occurance" remains O(n).
       *)
       IF NOT "Array.DInt.Is_Element"(dint_array := #dint_array, search_term := #search_term) THEN
           #"Array.DInt.First_Occurance" := -1;
           RETURN;
       END_IF;
       WHILE #dint_array[#_i] <> #search_term AND DINT_TO_UDINT(#_i) < #_length DO
           #_i += 1;
       END_WHILE;
   END_REGION


   REGION _name_
       #"Array.DInt.First_Occurance" := #_i;
   END_REGION
END_FUNCTION

FUNCTION "Array.DInt.Intersect_Exists" : Bool   // FC144, SCL
{ S7_Optimized_Access := 'TRUE' }
VERSION : 0.1
   VAR_INPUT
      "a" : Variant;   // should be array of dint, max 999
      "b" : Variant;   // should be array of dint, max 999
      null_value : DInt;
   END_VAR
   VAR_TEMP
      i : Int;
      j : Int;
      len_a : Struct
         as_udint : UDInt;
         as_int : Int;
      END_STRUCT;
      len_b : Struct
         as_udint : UDInt;
         as_int : Int;
      END_STRUCT;
      t_a : Array[0..#u_bound] of DInt;
      p_ret : Int;
      ret : Bool;
      t_b : Array[0..#u_bound] of DInt;
      status : Int;
   END_VAR
   VAR CONSTANT
      u_bound : Int := 999;
   END_VAR
BEGIN
   REGION "GET LENGHTS"
       #len_a.as_udint := CountOfElements(#a);
       #len_a.as_int := UDINT_TO_INT(#len_a.as_udint) - 1;
       #len_b.as_udint := CountOfElements(#b);
       #len_b.as_int := UDINT_TO_INT(#len_b.as_udint) - 1;
   END_REGION

   REGION "PERFORM MOVES"
       #status := MOVE_BLK_VARIANT(SRC := #a, COUNT := #len_a.as_udint, SRC_INDEX := 0, DEST_INDEX := 0, DEST => #t_a);
       #status := MOVE_BLK_VARIANT(SRC := #b, COUNT := #len_b.as_udint, SRC_INDEX := 0, DEST_INDEX := 0, DEST => #t_b);
   END_REGION


   REGION "SEARCH FOR ANY MATCHING ELEMENT"
       FOR #i := 0 TO #len_a.as_int DO

           REGION "SKIP NULL VALUES"
               IF #t_a[#i] = #null_value THEN
                   CONTINUE;
               END_IF;
           END_REGION

           REGION "INNER LOOP"
               FOR #j := 0 TO #len_b.as_int DO

                   REGION "SKIP NULL VALUES"
                       IF #t_b[#j] = #null_value THEN
                           CONTINUE;
                       END_IF;
                   END_REGION

                   REGION "SET RETURN VALUE ON MATCH"
                       IF #t_a[#i] = #t_b[#j] THEN
                           #ret := TRUE;
                           EXIT;
                       END_IF;
                   END_REGION

               END_FOR;
           END_REGION

           REGION "EXIT OUTTER LOOP IF MATCH FOUND"
               IF #ret THEN
                   EXIT;
               END_IF;
           END_REGION

       END_FOR;
   END_REGION

   REGION "RETURN"
       #"Array.DInt.Intersect_Exists" := #ret;
   END_REGION
END_FUNCTION

FUNCTION "Array.DInt.Intersect" : Void   // FC145, SCL
{ S7_Optimized_Access := 'TRUE' }
VERSION : 0.1
   VAR_INPUT
      "a" : Variant;   // should be array of dint, max 999
      "b" : Variant;   // should be array of dint, max 999
      null_value : DInt;
   END_VAR
   VAR_OUTPUT
      intersect_array : Variant;   // should be array of dint, max 999
   END_VAR
   VAR_TEMP
      i : Int;
      j : Int;
      len_a : Struct
         as_udint : UDInt;
         as_int : Int;
      END_STRUCT;
      len_b : Struct
         as_udint : UDInt;
         as_int : Int;
      END_STRUCT;
      t_a : Array[0..#u_bound] of DInt;
      p_ret : Int;
      ret : Array[0..#u_bound_double] of DInt;
      t_b : Array[0..#u_bound] of DInt;
      status : Int;
   END_VAR
   VAR CONSTANT
      u_bound : Int := 999;
      u_bound_double : Int := 1999;
   END_VAR
BEGIN
   REGION "GET LENGTHS"
       #len_a.as_udint := CountOfElements(#a);
       #len_a.as_int := UDINT_TO_INT(#len_a.as_udint) - 1;
       #len_b.as_udint := CountOfElements(#b);
       #len_b.as_int := UDINT_TO_INT(#len_b.as_udint) - 1;
   END_REGION

   REGION "MOVE"
       #status := MOVE_BLK_VARIANT(SRC := #a, COUNT := #len_a.as_udint, SRC_INDEX := 0, DEST_INDEX := 0, DEST => #t_a);
       #status := MOVE_BLK_VARIANT(SRC := #b, COUNT := #len_b.as_udint, SRC_INDEX := 0, DEST_INDEX := 0, DEST => #t_b);
   END_REGION

   REGION "FIND INTERSECT"
       FOR #i := 0 TO #len_a.as_int DO
           IF #t_a[#i] = #null_value THEN
               EXIT;
           END_IF;
           FOR #j := 0 TO #len_b.as_int DO
               IF #t_b[#j] = #null_value THEN
                   EXIT;
               END_IF;
               IF #t_a[#i] = #t_b[#j] THEN
                   #ret[#p_ret] := #t_a[#i];
                   #p_ret += 1;
                   EXIT;
               END_IF;
           END_FOR;
       END_FOR;
   END_REGION

   REGION "RETURN"
       #status := MOVE_BLK_VARIANT(SRC := #ret, COUNT := INT_TO_UDINT(#p_ret - 1), SRC_INDEX := 0, DEST_INDEX := 0, DEST => #intersect_array);
   END_REGION
END_FUNCTION

FUNCTION "Array.WString.Is_Element" : Bool   // FC207, SCL
{ S7_Optimized_Access := 'TRUE' }
VERSION : 0.1
   VAR_INPUT
      search_term : WString;
      search_array : Array[*] of WString[1];
   END_VAR
   VAR_TEMP
      _i : Int;
      _length_search_array : UDInt;
   END_VAR
BEGIN
   #_length_search_array := "Array.Any.Length"(#search_array);
   FOR #_i := 0 TO UDINT_TO_INT(#_length_search_array - 1) DO
       IF #search_term = #search_array[#_i] THEN
           #"Array.WString.Is_Element" := TRUE;
           RETURN;
       END_IF;
   END_FOR;
   #"Array.WString.Is_Element" := FALSE;
END_FUNCTION

FUNCTION "Array.Int.First_Occurance" : DInt   // FC220, SCL
{ S7_Optimized_Access := 'TRUE' }
VERSION : 0.1
   VAR_INPUT
      int_array : Array[*] of Int;
      search_term : Int;
   END_VAR
   VAR_TEMP
      _i : DInt;
      _length : UDInt;
   END_VAR
BEGIN
   REGION "NOTES"
       (* 
       This function returns the first occurance of the search term.
       This function meant for use with collapsed arrays.
       See "Array.Int.Collapse" for collapse functionality.
       *)
   END_REGION


   REGION "GET LENGTH OF INPUT ARRAY"
       #_length := "Array.Any.Length"(#int_array);
   END_REGION


   REGION "FIND FIRST SEARCH TERM, -1 IF NONE"
       (*
       Its worth noting that "Array.Int.Is_Element" could return the index of the search term
       as an output, saving the processor some work. 
       The rework is justified by increased encapsulation.
       The time complexity for "Array.Int.First_Occurance" remains O(n).
       *)
       IF NOT "Array.Int.Is_Element"(int_array := #int_array, search_term := #search_term) THEN
           #"Array.Int.First_Occurance" := -1;
           RETURN;
       END_IF;
       WHILE #int_array[#_i] <> #search_term AND DINT_TO_UDINT(#_i) < #_length DO
           #_i += 1;
       END_WHILE;
   END_REGION


   REGION _name_
       #"Array.Int.First_Occurance" := #_i;
   END_REGION
END_FUNCTION

FUNCTION "Array.WString.Fill" : Void   // FC243, SCL
{ S7_Optimized_Access := 'TRUE' }
VERSION : 0.1
   VAR_INPUT
      value : WString;
   END_VAR
   VAR_IN_OUT
      "array" : Array[*] of WString;
   END_VAR
   VAR_TEMP
      _length : Int;
      _i : Int;
   END_VAR
BEGIN
   #_length := UDINT_TO_INT("Array.Any.Length"(#array)) - 1;
   FOR #_i := 0 TO #_length DO
       #array[#_i] := #value;
   END_FOR;
   RETURN;
END_FUNCTION

FUNCTION "Array.WString.Search" : Int   // FC244, SCL
{ S7_Optimized_Access := 'TRUE' }
VERSION : 0.1
   VAR_INPUT
      "array" : Array[*] of WString;
      search_term : WString;
   END_VAR
   VAR_TEMP
      _i : Int;
      _length : Int;
   END_VAR
   // Ret_Val : index of search term. returns -1 if not found.
BEGIN
   REGION "SEARCH ARRAY"
       #_length := UDINT_TO_INT("Array.Any.Length"(#array)) - 1;
       FOR #_i := 0 TO #_length DO
           IF #array[#_i] <> #search_term THEN
               CONTINUE;
           END_IF;
           #"Array.WString.Search" := #_i;
           RETURN;
       END_FOR;
   END_REGION

   REGION "RETURN"
       #"Array.WString.Search" := "NULL_TOKEN";
       RETURN;
   END_REGION
END_FUNCTION

// folder: Utilities/Bool

FUNCTION "Bool.Animate" : USInt   // FC9, SCL
{ S7_Optimized_Access := 'TRUE' }
VERSION : 0.1
   VAR_INPUT
      true_color : USInt;
      false_color : USInt;
      evaluation_signal : Bool;
   END_VAR
   VAR_TEMP
      animate : USInt;
   END_VAR
BEGIN
   REGION "FALSE COLOR"
       IF NOT #evaluation_signal THEN
           #animate := #false_color;
       END_IF;
   END_REGION

   REGION "TRUE COLOR"
       IF #evaluation_signal THEN
           #animate := #true_color;
       END_IF;
   END_REGION

   REGION "FUNCTION RETURN"
       #"Bool.Animate" := #animate;
   END_REGION
END_FUNCTION

FUNCTION "Bool.Rising_Edge" : Bool   // FC177, SCL
{ S7_Optimized_Access := 'TRUE' }